PopupScreen "Comandos Perfiladores" 1280x714
   Button "Botón_6" at 630,585 size 88x33; TextOff 'Avance'
      on Press: SetTag("DB_OP.RC1", 52); SetBit("DB_OP.OP_SELMANU1")
      Visibility <- "MANU"
      Appearance <- "DB_OP.RC1"
   Button "Botón_7" at 630,630 size 88x33; TextOff 'Retroceso'
      on Press: SetTag("DB_OP.RC1", 53); SetBit("DB_OP.OP_SELMANU1")
      Visibility <- "MANU"
      Appearance <- "DB_OP.RC1"
   Button "Botón_8" at 731,585 size 88x33; TextOff 'Hacia Consigna'
      on Press: SetTag("DB_OP.RC1", 51); SetBit("DB_OP.OP_SELMANU1")
      Visibility <- "MANU"
      Appearance <- "DB_OP.RC1"
   Button "Botón_11" at 731,630 size 88x33; TextOff 'Freno'
      on Press: SetTag("DB_OP.RC1", 54); SetBit("DB_OP.OP_SELMANU1")
      Visibility <- "MANU"
      Appearance <- "DB_OP.RC1"
   Button "Botón_1" at 889,270 size 88x33; TextOff 'Avance'
      on Press: SetTag("DB_OP.RC1", 55); SetBit("DB_OP.OP_SELMANU1")
      Visibility <- "MANU"
      Appearance <- "DB_OP.RC1"
   Button "Botón_2" at 889,307 size 88x33; TextOff 'Retroceso'
      on Press: SetTag("DB_OP.RC1", 56); SetBit("DB_OP.OP_SELMANU1")
      Visibility <- "MANU"
      Appearance <- "DB_OP.RC1"
   IOField "Champ E/S_1" at 943,573 size 77x29; FormatPattern 9999999
      ProcessValue <- "DB_OP.COD1_VAL"
   IOField "Champ E/S" at 947,636 size 70x29; FormatPattern 9.9999
      ProcessValue <- "DB_OP.COD1_COEF"
   IOField "Champ E/S_0" at 943,601 size 77x29; FormatPattern 9999999
      ProcessValue <- "DB_OP.COD1_CONS"
   IOField "Champ E/S_2" at 1114,575 size 69x29; FormatPattern 9999999
      ProcessValue <- "DB_OP.COD1_INIT"
   TextField "Champ de texte_2" at 861,578 size 82x18; Text 'Posición / Position Réelle'
   TextField "Champ de texte" at 844,607 size 99x18; Text 'Consigna / Position Consigne'
   TextField "Champ de texte_0" at 851,641 size 92x18; Text 'Coef corrección / Coeff correction'
   IOField "Champ E/S_4" at 1114,640 size 69x29; FormatPattern 9999999
      ProcessValue <- "DB_OP.COD1_TARGET"
   TextField "Champ de texte_5" at 1044,612 size 62x18; Text 'Cota Paro / Côte Arrêt'
   TextField "Champ de texte_6" at 1052,645 size 50x18; Text 'Ventana / Fenetre'
   IOField "Champ E/S_5" at 1114,607 size 69x29; FormatPattern 9999999
      ProcessValue <- "DB_OP.COD1_ARRET"
   Button "Button" at 1045,578 size 60x23; TextOff 'OFFSET'; Authorization "Nivel 1"
      on Press: SetBit("DB_OP.COD1_CMD")
      Appearance <- "DB_OP.COD2_CMD"
   GraphicIOField "Campo ES gráfico_4" at 236,203 size 456x232; PictureList "Grupo 2 - Perfilador"
      ProcessValue <- "Alarma_Perfiladores"
   Polygon "Polígono_3" at 265,240 size 389x46
      Visibility <- "Perfiladores\Perfilador.PresenciaPieza"
   Rectangle "Rectángulo_2" at 874,227 size 118x128
      Visibility <- "MANU"
   Rectangle "Rectángulo_3" at 874,227 size 118x29
      Visibility <- "MANU"
   TextField "Campo de texto_1" at 900,231 size 66x18; Text 'Perfiladores'
      Visibility <- "MANU"
   Circle "Cercle_11" at 450,253 size 12x12
      Appearance <- "27S4"
   Circle "Cercle_12" at 413,405 size 12x12
      Appearance <- "29S7"
   Circle "Cercle_13" at 411,387 size 12x12
      Appearance <- "29S7"
   Circle "Cercle_14" at 515,384 size 12x12
      Appearance <- "23S4"
   Polygon "Polígono_1" at 248,269 size 17x19
      Appearance <- "36S70"
   TextField "Campo de texto_3" at 246,143 size 112x18; Text 'Sensores de Atasco'
   TextField "Campo de texto_4" at 613,454 size 141x18; Text '23S4 - Presión de Frenos'
   TextField "Campo de texto_5" at 414,107 size 101x18; Text 'Motor Perfilador 4'
   TextField "Campo de texto_6" at 684,429 size 101x18; Text 'Motor Perfilador 3'
   TextField "Campo de texto_7" at 159,441 size 101x18; Text 'Motor Perfilador 1'
   TextField "Campo de texto_8" at 147,165 size 101x18; Text 'Motor Perfilador 2'
   TextField "Campo de texto_9" at 140,188 size 64x46; Text '36S70 Barrera de Atascos'
   TextField "Campo de texto_10" at 557,500 size 197x18; Text 'M07 - Motor Ajuste de Profundidad'
   TextField "Campo de texto_11" at 202,476 size 119x18; Text '29S7 - Fin de Carrera'
   TextField "Campo de texto_13" at 320,502 size 53x18; Text 'Encóder'
   TextField "Campo de texto_14" at 118,363 size 81x46; Text '27S3 - Chapa en Entrada Perfilador'
   Circle "Cercle_2" at 236,274 size 12x12
      Appearance <- "27S3"
   Polyline "Línea poligonal_11" at 263,255 size 397x22
      Appearance <- "36S70"
   Polygon "Polígono_2" at 655,246 size 17x19
      Appearance <- "36S70"
   Rectangle "Rectángulo_6" at 613,555 size 222x128
      Visibility <- "MANU"
   Rectangle "Rectángulo_7" at 834,539 size 374x144
      Visibility <- "MANU"
   Rectangle "Rectángulo_8" at 613,539 size 595x29
      Visibility <- "MANU"
   TextField "Campo de texto_12" at 674,543 size 108x18; Text 'Ajuste Profundidad'
      Visibility <- "MANU"

PopupScreen "Comandos Cinta" 1280x714
   Button "Botón_6" at 630,585 size 88x33; TextOff 'Avance'
      on Press: SetTag("DB_OP.RC1", 52); SetBit("DB_OP.OP_SELMANU1")
      Visibility <- "MANU"
      Appearance <- "DB_OP.RC1"
   Button "Botón_7" at 630,630 size 88x33; TextOff 'Retroceso'
      on Press: SetTag("DB_OP.RC1", 53); SetBit("DB_OP.OP_SELMANU1")
      Visibility <- "MANU"
      Appearance <- "DB_OP.RC1"
   Button "Botón_8" at 731,585 size 88x33; TextOff 'Hacia Consigna'
      on Press: SetTag("DB_OP.RC1", 51); SetBit("DB_OP.OP_SELMANU1")
      Visibility <- "MANU"
      Appearance <- "DB_OP.RC1"
   Button "Botón_11" at 731,630 size 88x33; TextOff 'Freno'
      on Press: SetTag("DB_OP.RC1", 54); SetBit("DB_OP.OP_SELMANU1")
      Visibility <- "MANU"
      Appearance <- "DB_OP.RC1"
   Button "Botón_4" at 462,582 size 88x33; TextOff 'Avance'
      on Press: SetTag("DB_OP.RC2", 91); SetBit("DB_OP.OP_SELMANU2")
      Visibility <- "MANU"
      Appearance <- "DB_OP.RC2"
   Button "Botón_5" at 462,619 size 88x33; TextOff 'Retroceso'
      on Press: SetTag("DB_OP.RC2", 92); SetBit("DB_OP.OP_SELMANU2")
      Visibility <- "MANU"
      Appearance <- "DB_OP.RC2"
   IOField "Champ E/S_1" at 943,573 size 77x29; FormatPattern 9999999
      ProcessValue <- "DB_OP.COD2_VAL"
   IOField "Champ E/S" at 947,636 size 70x29; FormatPattern 9.9999
      ProcessValue <- "DB_OP.COD2_COEF"
   IOField "Champ E/S_0" at 943,601 size 77x29; FormatPattern 9999999
      ProcessValue <- "DB_OP.COD2_CONS"
   IOField "Champ E/S_2" at 1114,575 size 69x29; FormatPattern 9999999
      ProcessValue <- "DB_OP.COD2_INIT"
   TextField "Champ de texte_2" at 861,578 size 82x18; Text 'Posición / Position Réelle'
   TextField "Champ de texte" at 844,607 size 99x18; Text 'Consigna / Position Consigne'
   TextField "Champ de texte_0" at 851,641 size 92x18; Text 'Coef corrección / Coeff correction'
   IOField "Champ E/S_4" at 1114,640 size 69x29; FormatPattern 9999999
      ProcessValue <- "DB_OP.COD2_TARGET"
   TextField "Champ de texte_5" at 1044,612 size 62x18; Text 'Cota Paro / Côte Arrêt'
   TextField "Champ de texte_6" at 1052,645 size 50x18; Text 'Ventana / Fenetre'
   IOField "Champ E/S_5" at 1114,607 size 69x29; FormatPattern 9999999
      ProcessValue <- "DB_OP.COD2_ARRET"
   Button "Button" at 1045,578 size 60x23; TextOff 'OFFSET'; Authorization "Nivel 1"
      on Press: SetBit("DB_OP.COD2_CMD")
      Appearance <- "DB_OP.COD2_CMD"
   GraphicIOField "Campo ES gráfico_1" at 290,222 size 647x180; PictureList "Grupo 2 - Cinta"
      ProcessValue <- "Alarma_Cinta"
   Rectangle "Rectángulo_1" at 613,555 size 222x128
      Visibility <- "MANU"
   Rectangle "Rectángulo_2" at 448,539 size 118x128
      Visibility <- "MANU"
   Rectangle "Rectángulo_3" at 448,539 size 118x29
      Visibility <- "MANU"
   TextField "Campo de texto_1" at 474,543 size 31x18; Text 'Cinta'
      Visibility <- "MANU"
   Rectangle "Rectángulo_6" at 834,539 size 374x144
      Visibility <- "MANU"
   Rectangle "Rectángulo_7" at 613,539 size 595x29
      Visibility <- "MANU"
   TextField "Campo de texto_12" at 642,543 size 108x18; Text 'Ajuste Profundidad'
      Visibility <- "MANU"
   Circle "Cercle_1" at 325,248 size 12x12
      Appearance <- "27S4"
   Circle "Cercle_14" at 909,220 size 12x12
      Appearance <- "29S1"
   Circle "Cercle_15" at 909,234 size 12x12
      Appearance <- "29S2"
   Circle "Cercle_11" at 826,289 size 12x12
      Appearance <- "25S2"
   Circle "Cercle" at 911,284 size 12x12
      Appearance <- "29S3"
   TextField "Campo de texto_22" at 109,219 size 183x18; Text '27S4 - Chapa en Salida Perfilador'
   TextField "Campo de texto_23" at 624,433 size 179x18; Text 'M07 - Motor Ajuste Profundidad'
   TextField "Campo de texto_24" at 987,328 size 126x18; Text '25S2 - Bajar Velocidad'
   TextField "Campo de texto_25" at 512,385 size 223x18; Text '29S3 - Presencia de Chapa en Formador'
   TextField "Campo de texto_31" at 616,197 size 166x18; Text 'M08 - Motor Transporte Cinta'
   TextField "Campo de texto_32" at 667,130 size 145x18; Text '29S1 - Avance Bloqueado'
   TextField "Campo de texto_33" at 647,164 size 165x18; Text '29S2 - Avance Desbloqueado'
   Polygon "Polígono_4" at 351,252 size 385x62
      Visibility <- "Cinta\Cinta.PresenciaPieza"

PopupScreen "Comandos Descargador" 1280x714
   GraphicView "Visor de gráficos_1" at 134,166 size 538x272; Picture "Rolos 3"
   Rectangle "Rectángulo_9" at 811,197 size 118x128
      Visibility <- "MANU"
   Rectangle "Rectángulo_8" at 811,197 size 118x29
      Visibility <- "MANU"
   TextField "Campo de texto_3" at 854,201 size 32x18; Text 'Rolos'
      Visibility <- "MANU"
   Button "Botón_29" at 826,241 size 88x33; TextOff 'Avance'
      on Press: SetTag("DB_OP.RC1", 41); SetBit("DB_OP.OP_SELMANU1")
      Visibility <- "MANU"
      Appearance <- "DB_OP.RC1"
   Button "Botón_30" at 826,279 size 88x33; TextOff 'Retroceso'
      on Press: SetTag("DB_OP.RC1", 42); SetBit("DB_OP.OP_SELMANU1")
      Visibility <- "MANU"
      Appearance <- "DB_OP.RC1"
   TextField "Campo de texto_7" at 303,476 size 104x32; Text '27S3 - Chapa en Entrada Perfilador'
   Circle "Cercle_10" at 201,328 size 12x12
      Appearance <- "27S3"
   Circle "Cercle_13" at 349,283 size 12x12
      Appearance <- "26S8"
   TextField "Campo de texto_11" at 455,437 size 114x32; Text '26S8 - Chapa en Transporte de Rolos'

screen "eProC - 01 Araña" 1280x768, template "Template"
   Polygon "Polígono_3" at 343,318 size 325x50
      Visibility <- "Araña\Araña.PresenciaPieza"
   Rectangle "Rectángulo_7" at 989,250 size 248x208
      Visibility <- "MANU"
   Rectangle "Rectángulo_12" at 989,246 size 248x29
      Visibility <- "MANU"
   Rectangle "Rectángulo_9" at 843,563 size 118x128
      Visibility <- "MANU"
   Rectangle "Rectángulo_8" at 843,563 size 118x29
      Visibility <- "MANU"
   TextField "Campo de texto_3" at 870,567 size 64x18; Text 'Transporte'
      Visibility <- "MANU"
   TextField "Campo de texto_11" at 1010,252 size 66x18; Text 'Aire Tulipas'
      Visibility <- "MANU"
   Button "Botón_4" at 859,607 size 88x33; TextOff 'Avance'
      on Press: SetTag("DB_OP.RC1", 11); SetBit("DB_OP.OP_SELMANU1")
      Visibility <- "MANU"
      Appearance <- "DB_OP.RC1"
   Button "Botón_5" at 859,645 size 88x33; TextOff 'Retroceso'
      on Press: SetTag("DB_OP.RC1", 12); SetBit("DB_OP.OP_SELMANU1")
      Visibility <- "MANU"
      Appearance <- "DB_OP.RC1"
   Button "Botón_10" at 1065,290 size 72x33; TextOff 'Activar'
      on Press: SetTag("DB_OP.RC1", 20); SetBit("DB_OP.OP_SELMANU1")
      Visibility <- "MANU"
      Appearance <- "DB_OP.RC1"
   Button "Botón_17" at 1145,290 size 72x33; TextOff 'Desactivar'
      on Press: SetTag("DB_OP.RC1", 21); SetBit("DB_OP.OP_SELMANU1")
      Visibility <- "MANU"
      Appearance <- "DB_OP.RC1"
   TextField "Campo de texto_12" at 1010,296 size 37x18; Text 'Todas'
      Visibility <- "MANU"
   Button "Botón_1" at 1065,336 size 72x33; TextOff 'Activar'
      on Press: SetTag("DB_OP.RC1", 32); SetBit("DB_OP.OP_SELMANU1")
      Visibility <- "MANU"
      Appearance <- "DB_OP.RC1"
   Button "Botón_23" at 1065,373 size 72x33; TextOff 'Activar'
      on Press: SetTag("DB_OP.RC1", 34); SetBit("DB_OP.OP_SELMANU1")
      Visibility <- "MANU"
      Appearance <- "DB_OP.RC1"
   Button "Botón_24" at 1065,411 size 72x33; TextOff 'Activar'
      on Press: SetTag("DB_OP.RC1", 36); SetBit("DB_OP.OP_SELMANU1")
      Visibility <- "MANU"
      Appearance <- "DB_OP.RC1"
   Button "Botón_26" at 1145,336 size 72x33; TextOff 'Desactivar'
      on Press: SetTag("DB_OP.RC1", 33); SetBit("DB_OP.OP_SELMANU1")
      Visibility <- "MANU"
      Appearance <- "DB_OP.RC1"
   Button "Botón_27" at 1145,373 size 72x33; TextOff 'Desactivar'
      on Press: SetTag("DB_OP.RC1", 35); SetBit("DB_OP.OP_SELMANU1")
      Visibility <- "MANU"
      Appearance <- "DB_OP.RC1"
   Button "Botón_28" at 1145,411 size 72x33; TextOff 'Desactivar'
      on Press: SetTag("DB_OP.RC1", 37); SetBit("DB_OP.OP_SELMANU1")
      Visibility <- "MANU"
      Appearance <- "DB_OP.RC1"
   TextField "Campo de texto_2" at 1008,343 size 48x18; Text 'Grupo 1'
      Visibility <- "MANU"
   TextField "Campo de texto_1" at 1008,381 size 48x18; Text 'Grupo 2'
      Visibility <- "MANU"
   TextField "Campo de texto_5" at 1008,419 size 48x18; Text 'Grupo 3'
      Visibility <- "MANU"
   Rectangle "Rectángulo_1" at 989,483 size 248x208
      Visibility <- "MANU"
   Rectangle "Rectángulo_2" at 989,479 size 248x29
      Visibility <- "MANU"
   TextField "Campo de texto_13" at 1010,485 size 74x18; Text 'Vacío Tulipas'
      Visibility <- "MANU"
   TextField "Campo de texto_14" at 1010,529 size 37x18; Text 'Todas'
      Visibility <- "MANU"
   TextField "Campo de texto_15" at 1008,576 size 48x18; Text 'Grupo 1'
      Visibility <- "MANU"
   TextField "Campo de texto_16" at 1008,614 size 48x18; Text 'Grupo 2'
      Visibility <- "MANU"
   TextField "Campo de texto_17" at 1008,652 size 48x18; Text 'Grupo 3'
      Visibility <- "MANU"
   Button "Botón_21" at 1065,523 size 72x33; TextOff 'Activar'
      on Press: SetTag("DB_OP.RC1", 30); SetBit("DB_OP.OP_SELMANU1")
      Visibility <- "MANU"
      Appearance <- "DB_OP.RC1"
   Button "Botón_25" at 1145,523 size 72x33; TextOff 'Desactivar'
      on Press: SetTag("DB_OP.RC1", 31); SetBit("DB_OP.OP_SELMANU1")
      Visibility <- "MANU"
      Appearance <- "DB_OP.RC1"
   Button "Botón_14" at 1065,569 size 72x33; TextOff 'Activar'
      on Press: SetTag("DB_OP.RC1", 22); SetBit("DB_OP.OP_SELMANU1")
      Visibility <- "MANU"
      Appearance <- "DB_OP.RC1"
   Button "Botón_15" at 1065,606 size 72x33; TextOff 'Activar'
      on Press: SetTag("DB_OP.RC1", 24); SetBit("DB_OP.OP_SELMANU1")
      Visibility <- "MANU"
      Appearance <- "DB_OP.RC1"
   Button "Botón_16" at 1065,644 size 72x33; TextOff 'Activar'
      on Press: SetTag("DB_OP.RC1", 26); SetBit("DB_OP.OP_SELMANU1")
      Visibility <- "MANU"
      Appearance <- "DB_OP.RC1"
   Button "Botón_18" at 1145,569 size 72x33; TextOff 'Desactivar'
      on Press: SetTag("DB_OP.RC1", 23); SetBit("DB_OP.OP_SELMANU1")
      Visibility <- "MANU"
      Appearance <- "DB_OP.RC1"
   Button "Botón_19" at 1145,606 size 72x33; TextOff 'Desactivar'
      on Press: SetTag("DB_OP.RC1", 25); SetBit("DB_OP.OP_SELMANU1")
      Visibility <- "MANU"
      Appearance <- "DB_OP.RC1"
   Button "Botón_20" at 1145,644 size 72x33; TextOff 'Desactivar'
      on Press: SetTag("DB_OP.RC1", 27); SetBit("DB_OP.OP_SELMANU1")
      Visibility <- "MANU"
      Appearance <- "DB_OP.RC1"
   Rectangle "Rectángulo_10" at 988,26 size 248x201
      Visibility <- "MANU"
   Button "Botón_6" at 1012,65 size 202x33; TextOff 'Subir (Pistón Superior)'
      on Press: SetTag("DB_OP.RC1", 16); SetBit("DB_OP.OP_SELMANU1")
      Visibility <- "MANU"
      Appearance <- "DB_OP.RC1"
   Button "Botón_7" at 1012,103 size 202x33; TextOff 'Bajar (Pistón Superior)'
      on Press: SetTag("DB_OP.RC1", 15); SetBit("DB_OP.OP_SELMANU1")
      Visibility <- "MANU"
      Appearance <- "DB_OP.RC1"
   Button "Botón_8" at 1012,179 size 202x33; TextOff 'Bajar (Pistón Inferior)'
      on Press: SetTag("DB_OP.RC1", 13); SetBit("DB_OP.OP_SELMANU1")
      Visibility <- "MANU"
      Appearance <- "DB_OP.RC1"
   Button "Botón_9" at 1012,141 size 202x33; TextOff 'Subir (Pistón Inferior)'
      on Press: SetTag("DB_OP.RC1", 14); SetBit("DB_OP.OP_SELMANU1")
      Visibility <- "MANU"
      Appearance <- "DB_OP.RC1"
   Rectangle "Rectángulo_11" at 988,26 size 248x29
      Visibility <- "MANU"
   TextField "Campo de texto_7" at 1056,30 size 110x18; Text 'Movimiento Vertical'
      Visibility <- "MANU"
   GraphicIOField "Campo ES gráfico_1" at 295,98 size 460x334; PictureList "Araña"
      ProcessValue <- "Alarma_Araña"
   Button "Botón_2" at 453,467 size 144x49; TextOff 'Inicializar'
      on Press: SetBit("Comando_Inicializar_Araña")
      Visibility <- "MANU"
   Group "Group" at 428,460 size 189x68
   TextField "Campo de texto_8" at 61,77 size 35x18; Text 'Araña'
   TextField "Campo de texto_18" at 61,98 size 12x18; Text 'A'
   IOField "Champ E/S_8" at 98,95 size 54x25; FormatPattern 9999999
      Appearance <- "Araña\Araña.PresenciaPieza"
      ProcessValue <- "Araña\Araña.A"
   IOField "Champ E/S_9" at 98,115 size 54x25; FormatPattern 9999999
      Appearance <- "Araña\Araña.PresenciaPieza"
      ProcessValue <- "Araña\Araña.B"
   IOField "Champ E/S_10" at 98,136 size 54x24; FormatPattern 9999999
      Appearance <- "Araña\Araña.PresenciaPieza"
      ProcessValue <- "Araña\Araña.C"
   IOField "Champ E/S_11" at 98,155 size 54x25; FormatPattern 9999999
      Appearance <- "Araña\Araña.PresenciaPieza"
      ProcessValue <- "Araña\Araña.D"
   TextField "Campo de texto_29" at 62,116 size 11x18; Text 'B'
   TextField "Campo de texto_30" at 62,136 size 11x18; Text 'C'
   TextField "Campo de texto_31" at 62,156 size 12x18; Text 'D'
   Button "Botón_3" at 45,40 size 128x33; TextOff 'Borrar Pieza'
      on Click: ResetBit("Araña\Araña.PresenciaPieza")
      Visibility <- "Araña\Araña.PresenciaPieza"
   Button "Botón_12" at 45,340 size 128x33; TextOff 'Transferir Datos'
      on Click: SetBit("Forz_Transf1")
      Visibility <- "Perfiladores\Perfilador.PresenciaPieza"
   Button "Template_Plantilla_Botón_3" at 1,688 size 130x29; TextOff 'ARAÑA'
   Button "Plantilla_Botón_1" at 1,715 size 130x53; TextOff 'PRINCIPAL'
      on Click: ActivateScreen("eProC - Principal", 0)
   Button "Template_Plantilla_Bouton_2" at 1085,715 size 193x53; TextOff 'ALARMAS / DEFAUT'
      on Press: ActivateScreen("eProC - Alarmas", 0)
      Visibility <- "DB_OP.P_DEFAUT"
   Circle "Cercle_11" at 494,226 size 10x10
      Appearance <- "25S8"
   Circle "Cercle_12" at 495,183 size 10x10
      Appearance <- "25S7"
   Circle "Cercle_0" at 494,247 size 10x10
      Appearance <- "25S4"
   Circle "Cercle_1" at 534,134 size 10x10
      Appearance <- "25S3"
   Circle "Cercle_2" at 538,186 size 10x10
      Appearance <- "25S5"
   TextField "Campo de texto_6" at 645,56 size 186x22; Text '25S3 - Fin de Carrera Arriba'
   TextField "Campo de texto_9" at 620,126 size 186x22; Text '25S5 - Fin de Carrera Abajo'
   TextField "Campo de texto_19" at 218,103 size 174x22; Text '25S7 - Pistón 2 Expandido'
   TextField "Campo de texto_20" at 220,139 size 169x22; Text '25S8 - Pistón 2 Contraído'
   TextField "Campo de texto_21" at 220,198 size 169x22; Text '25S4 - Pistón 1 Contraído'
   TextField "Campo de texto_22" at 297,228 size 132x22; Text '25S6 - Araña Abajo'
   Circle "Cercle_5" at 457,251 size 10x10
      Appearance <- "25S6"
   Circle "Cercle" at 476,339 size 10x10
      Appearance <- "26S1"
   TextField "Campo de texto_23" at 183,430 size 248x22; Text '26S1 - Tulipas Apoyadas en la Chapa'
   TextField "Campo de texto_24" at 768,228 size 151x22; Text '26S5 - Bajar Velocidad'
   TextField "Campo de texto_25" at 763,204 size 210x22; Text '26S3 - En Posición de Descarga'
   TextField "Campo de texto_26" at 773,293 size 206x58; Text 'M03 - Motor Transporte Araña KM02.1 -> Hacia Rolos KM02.2 -> Hacia Almacenes'
   TextField "Campo de texto_27" at 785,393 size 151x22; Text '26S4 - Bajar Velocidad'
   TextField "Campo de texto_28" at 787,418 size 187x22; Text '26S2 - En Posición de Carga'
   Circle "Cercle_4" at 701,406 size 10x10
      Appearance <- "26S2"
   Circle "Cercle_6" at 696,382 size 10x10
      Appearance <- "26S4"
   Circle "Cercle_7" at 681,214 size 10x10
      Appearance <- "26S5"
   Circle "Cercle_8" at 676,191 size 10x10
      Appearance <- "26S3"
   Rectangle "Rectángulo_3" at 428,460 size 189x68
      Visibility <- "Araña_Inicializada"
   TextField "Campo de texto_4" at 442,481 size 159x22; Text 'Araña en Posición Inicial'
      Visibility <- "Araña_Inicializada"
   TextField "Campo de texto_142" at 62,178 size 17x18; Text 'F1'
   IOField "Champ E/S_134" at 102,175 size 51x25; FormatPattern s999999
      Appearance <- "Araña\Araña.PresenciaPieza"
      ProcessValue <- "Araña\Araña.F1"
   IOField "Champ E/S_135" at 102,195 size 51x25; FormatPattern s999999
      Appearance <- "Araña\Araña.PresenciaPieza"
      ProcessValue <- "Araña\Araña.F2"
   IOField "Champ E/S_136" at 102,216 size 51x24; FormatPattern s999999
      Appearance <- "Araña\Araña.PresenciaPieza"
      ProcessValue <- "Araña\Araña.F3"
   IOField "Champ E/S_137" at 102,235 size 51x25; FormatPattern s999999
      Appearance <- "Araña\Araña.PresenciaPieza"
      ProcessValue <- "Araña\Araña.F4"
   TextField "Campo de texto_143" at 62,197 size 17x18; Text 'F2'
   TextField "Campo de texto_144" at 62,217 size 17x18; Text 'F3'
   TextField "Campo de texto_145" at 62,237 size 17x18; Text 'F4'
   TextField "Campo de texto_146" at 62,258 size 35x18; Text 'PL1-1'
   IOField "Champ E/S_138" at 102,255 size 51x25; FormatPattern s999999
      Appearance <- "Araña\Araña.PresenciaPieza"
      ProcessValue <- "Araña\Araña.PL1_1"
   IOField "Champ E/S_139" at 102,275 size 51x25; FormatPattern s999999
      Appearance <- "Araña\Araña.PresenciaPieza"
      ProcessValue <- "Araña\Araña.PL1_2"
   IOField "Champ E/S_140" at 102,296 size 51x24; FormatPattern s999999
      Appearance <- "Araña\Araña.PresenciaPieza"
      ProcessValue <- "Araña\Araña.PL2_1"
   IOField "Champ E/S_141" at 102,315 size 51x25; FormatPattern s999999
      Appearance <- "Araña\Araña.PresenciaPieza"
      ProcessValue <- "Araña\Araña.PL2_2"
   TextField "Campo de texto_147" at 62,278 size 35x18; Text 'PL1-2'
   TextField "Campo de texto_148" at 62,299 size 35x18; Text 'PL2-1'
   TextField "Campo de texto_149" at 62,318 size 35x18; Text 'PL2-2'

screen "eProC - 02 Rolos" 1280x768, template "Template"
   GraphicIOField "Campo ES gráfico_4" at 286,166 size 538x272; PictureList "Rolos"
      ProcessValue <- "Alarma_Perfiladores"
   Polygon "Polígono_3" at 336,215 size 385x136
      Visibility <- "Rolos\Rolos.PresenciaPieza"
   Rectangle "Rectángulo_9" at 963,197 size 118x128
      Visibility <- "MANU"
   Rectangle "Rectángulo_8" at 963,197 size 118x29
      Visibility <- "MANU"
   TextField "Campo de texto_3" at 1006,201 size 32x18; Text 'Rolos'
      Visibility <- "MANU"
   Button "Botón_29" at 978,241 size 88x33; TextOff 'Avance'
      on Press: SetTag("DB_OP.RC1", 41); SetBit("DB_OP.OP_SELMANU1")
      Visibility <- "MANU"
      Appearance <- "DB_OP.RC1"
   Button "Botón_30" at 978,279 size 88x33; TextOff 'Retroceso'
      on Press: SetTag("DB_OP.RC1", 42); SetBit("DB_OP.OP_SELMANU1")
      Visibility <- "MANU"
      Appearance <- "DB_OP.RC1"
   TextField "Campo de texto_7" at 455,476 size 124x40; Text '27S3 - Chapa en Entrada Perfilador'
   Circle "Cercle_10" at 353,328 size 12x12
      Appearance <- "27S3"
   Circle "Cercle_13" at 613,248 size 12x12
      Appearance <- "26S8"
   TextField "Campo de texto_11" at 719,402 size 137x40; Text '26S8 - Chapa en Transporte de Rolos'
   TextField "Campo de texto_10" at 61,77 size 32x18; Text 'Rolos'
   TextField "Campo de texto_20" at 61,99 size 12x18; Text 'A'
   IOField "Champ E/S_12" at 96,95 size 54x25; FormatPattern 9999999
      Appearance <- "Rolos\Rolos.PresenciaPieza"
      ProcessValue <- "Rolos\Rolos.A"
   IOField "Champ E/S_13" at 96,115 size 54x25; FormatPattern 9999999
      Appearance <- "Rolos\Rolos.PresenciaPieza"
      ProcessValue <- "Rolos\Rolos.B"
   IOField "Champ E/S_14" at 96,136 size 54x24; FormatPattern 9999999
      Appearance <- "Rolos\Rolos.PresenciaPieza"
      ProcessValue <- "Rolos\Rolos.C"
   IOField "Champ E/S_15" at 96,155 size 54x25; FormatPattern 9999999
      Appearance <- "Rolos\Rolos.PresenciaPieza"
      ProcessValue <- "Rolos\Rolos.D"
   TextField "Campo de texto_21" at 61,117 size 11x18; Text 'B'
   TextField "Campo de texto_22" at 61,137 size 11x18; Text 'C'
   TextField "Campo de texto_23" at 61,157 size 12x18; Text 'D'
   Button "Botón_9" at 45,40 size 126x33; TextOff 'Borrar Pieza'
      on Click: ResetBit("Rolos\Rolos.PresenciaPieza")
      Visibility <- "Rolos\Rolos.PresenciaPieza"
   Button "Botón_4" at 45,340 size 128x33; TextOff 'Transferir Datos'
      on Click: SetBit("Forz_Transf2")
      Visibility <- "Perfiladores\Perfilador.PresenciaPieza"
   Button "Template_Plantilla_Botón_3" at 1,688 size 130x29; TextOff 'ROLOS'
   Button "Plantilla_Botón_1" at 1,715 size 130x53; TextOff 'PRINCIPAL'
      on Click: ActivateScreen("eProC - Principal", 0)
   Button "Template_Plantilla_Bouton_2" at 1085,715 size 193x53; TextOff 'ALARMAS / DEFAUT'
      on Press: ActivateScreen("eProC - Alarmas", 0)
      Visibility <- "DB_OP.P_DEFAUT"
   TextField "Campo de texto_134" at 62,178 size 17x18; Text 'F1'
   IOField "Champ E/S_126" at 102,175 size 51x25; FormatPattern s999999
      Appearance <- "Rolos\Rolos.PresenciaPieza"
      ProcessValue <- "Rolos\Rolos.F1"
   IOField "Champ E/S_127" at 102,195 size 51x25; FormatPattern s999999
      Appearance <- "Rolos\Rolos.PresenciaPieza"
      ProcessValue <- "Rolos\Rolos.F2"
   IOField "Champ E/S_128" at 102,216 size 51x24; FormatPattern s999999
      Appearance <- "Rolos\Rolos.PresenciaPieza"
      ProcessValue <- "Rolos\Rolos.F3"
   IOField "Champ E/S_129" at 102,235 size 51x25; FormatPattern s999999
      Appearance <- "Rolos\Rolos.PresenciaPieza"
      ProcessValue <- "Rolos\Rolos.F4"
   TextField "Campo de texto_135" at 62,197 size 17x18; Text 'F2'
   TextField "Campo de texto_136" at 62,217 size 17x18; Text 'F3'
   TextField "Campo de texto_137" at 62,237 size 17x18; Text 'F4'
   TextField "Campo de texto_138" at 62,258 size 35x18; Text 'PL1-1'
   IOField "Champ E/S_130" at 102,255 size 51x25; FormatPattern s999999
      Appearance <- "Rolos\Rolos.PresenciaPieza"
      ProcessValue <- "Rolos\Rolos.PL1_1"
   IOField "Champ E/S_131" at 102,275 size 51x25; FormatPattern s999999
      Appearance <- "Rolos\Rolos.PresenciaPieza"
      ProcessValue <- "Rolos\Rolos.PL1_2"
   IOField "Champ E/S_132" at 102,296 size 51x24; FormatPattern s999999
      Appearance <- "Rolos\Rolos.PresenciaPieza"
      ProcessValue <- "Rolos\Rolos.PL2_1"
   IOField "Champ E/S_133" at 102,315 size 51x25; FormatPattern s999999
      Appearance <- "Rolos\Rolos.PresenciaPieza"
      ProcessValue <- "Rolos\Rolos.PL2_2"
   TextField "Campo de texto_139" at 62,278 size 35x18; Text 'PL1-2'
   TextField "Campo de texto_140" at 62,299 size 35x18; Text 'PL2-1'
   TextField "Campo de texto_141" at 62,318 size 35x18; Text 'PL2-2'

screen "eProC - 00 Almacenes" 1280x768, template "Template"
   Rectangle "Rectángulo_9" at 1020,194 size 118x128
      Visibility <- "MANU"
   Rectangle "Rectángulo_8" at 1020,194 size 118x29
      Visibility <- "MANU"
   TextField "Campo de texto_3" at 1036,198 size 86x18; Text 'Intercambiador'
      Visibility <- "MANU"
   Button "Botón_1" at 1035,238 size 88x33; TextOff 'Avance'
      on Press: SetTag("DB_OP.RC1", 1); SetBit("DB_OP.OP_SELMANU1")
      Visibility <- "MANU"
      Appearance <- "DB_OP.RC1"
   Button "Botón_2" at 1035,276 size 88x33; TextOff 'Retroceso'
      on Press: SetTag("DB_OP.RC1", 2); SetBit("DB_OP.OP_SELMANU1")
      Visibility <- "MANU"
      Appearance <- "DB_OP.RC1"
   TextField "Campo de texto_2" at 95,341 size 267x22; Text '26S7 - Almacén 2 en puesto de Trabajo'
   TextField "Campo de texto_4" at 175,412 size 260x22; Text '26S6 - Almacén 2 en puesto de Espera'
   GraphicIOField "Campo ES gráfico_2" at 480,113 size 396x294; PictureList "Grupo 1 - Almacén A"
      ProcessValue <- "26S7"
   GraphicIOField "Campo ES gráfico_1" at 480,113 size 396x294; PictureList "Grupo 1 - Almacén B"
      ProcessValue <- "26S7"
      Visibility <- "Alarma_Almacenes"
   Circle "Cercle_2" at 486,298 size 14x14
      Appearance <- "26S7"
   TextField "Campo de texto_6" at 132,470 size 286x22; Text 'M01 - Motor Intercambiador de Almacenes'
   Circle "Cercle_1" at 565,354 size 14x14
      Appearance <- "26S6"
   Polyline "Línea poligonal_11" at 542,162 size 264x133
      Appearance <- "36S10"
   TextField "Campo de texto_1" at 114,231 size 251x22; Text '36S10 - Barrera Seguridad Almacenes'
   Button "Botón_4" at 806,409 size 144x49; TextOff 'Habilitar'
      on Press: SetBit("Hab_Almacenes")
   Rectangle "Rectángulo_3" at 781,402 size 189x68
      Visibility <- "Enclavamiento"
   TextField "Campo de texto_5" at 800,423 size 148x22; Text 'Almacenes Habilitados'
      Visibility <- "Enclavamiento"
   Polygon "Polígono_2" at 800,152 size 20x12
      Appearance <- "36S10"
   Polygon "Polígono_1" at 528,288 size 20x12
      Appearance <- "36S10"
   Button "Template_Plantilla_Botón_3" at 1,688 size 130x29; TextOff 'ALMACENES'
   Button "Plantilla_Botón_1" at 1,715 size 130x53; TextOff 'PRINCIPAL'
      on Click: ActivateScreen("eProC - Principal", 0)
   Button "Template_Plantilla_Bouton_2" at 1085,715 size 193x53; TextOff 'ALARMAS / DEFAUT'
      on Press: ActivateScreen("eProC - Alarmas", 0)
      Visibility <- "DB_OP.P_DEFAUT"

screen "eProC - 03 Perfilador" 1280x768, template "Template"
   GraphicIOField "Campo ES gráfico_4" at 412,155 size 456x232; PictureList "Grupo 2 - Perfilador"
      ProcessValue <- "Alarma_Perfiladores"
   Polygon "Polígono_3" at 441,192 size 389x46
      Visibility <- "Perfiladores\Perfilador.PresenciaPieza"
   Rectangle "Rectángulo_2" at 987,531 size 118x144
      Visibility <- "MANU"
   Rectangle "Rectángulo_3" at 987,531 size 118x29
      Visibility <- "MANU"
   TextField "Campo de texto_1" at 1013,535 size 66x18; Text 'Perfiladores'
      Visibility <- "MANU"
   Circle "Cercle_11" at 458,214 size 12x12
      Appearance <- "Sensor 1"
   Circle "Cercle_13" at 587,339 size 12x12
      Appearance <- "29S6"
   Circle "Cercle_14" at 635,352 size 12x12
      Appearance <- "23S4"
   Polygon "Polígono_1" at 424,221 size 17x19
      Appearance <- "36S70"
   TextField "Campo de texto_3" at 406,92 size 134x22; Text 'Sensores de Atasco'
   TextField "Campo de texto_4" at 691,478 size 168x22; Text '23S4 - Presión de Frenos'
   TextField "Campo de texto_5" at 574,57 size 120x22; Text 'Motor Perfilador 4'
   TextField "Campo de texto_6" at 860,381 size 120x22; Text 'Motor Perfilador 3'
   TextField "Campo de texto_7" at 313,391 size 120x22; Text 'Motor Perfilador 1'
   TextField "Campo de texto_8" at 303,116 size 120x22; Text 'Motor Perfilador 2'
   TextField "Campo de texto_9" at 331,141 size 79x58; Text '36S70 Barrera de Atascos'
   TextField "Campo de texto_10" at 733,452 size 234x22; Text 'M07 - Motor Ajuste de Profundidad'
   TextField "Campo de texto_11" at 252,426 size 245x22; Text '29S6 - Fin de Carrera Hacia Adelante'
   TextField "Campo de texto_13" at 496,454 size 62x22; Text 'Encóder'
   TextField "Campo de texto_14" at 278,312 size 98x58; Text '27S3 - Chapa en Entrada Perfilador'
   Circle "Cercle_2" at 412,226 size 12x12
      Appearance <- "27S3"
   Polyline "Línea poligonal_11" at 439,207 size 397x22
      Appearance <- "36S70"
   Polygon "Polígono_2" at 831,198 size 17x19
      Appearance <- "36S70"
   Rectangle "Rectángulo_6" at 357,547 size 222x128
      Visibility <- "MANU"
   Rectangle "Rectángulo_8" at 357,531 size 222x29
      Visibility <- "MANU"
   TextField "Campo de texto_12" at 418,535 size 108x18; Text 'Ajuste Profundidad'
      Visibility <- "MANU"
   TextField "Campo de texto_2" at 61,77 size 54x18; Text 'Perfilador'
   TextField "Campo de texto_24" at 61,99 size 12x18; Text 'A'
   IOField "Champ E/S_16" at 100,95 size 53x25; FormatPattern 9999999
      Appearance <- "Perfiladores\Perfilador.PresenciaPieza"
      ProcessValue <- "Perfiladores\Perfilador.A"
   IOField "Champ E/S_17" at 100,115 size 53x25; FormatPattern 9999999
      Appearance <- "Perfiladores\Perfilador.PresenciaPieza"
      ProcessValue <- "Perfiladores\Perfilador.B"
   IOField "Champ E/S_18" at 100,136 size 53x24; FormatPattern 9999999
      Appearance <- "Perfiladores\Perfilador.PresenciaPieza"
      ProcessValue <- "Perfiladores\Perfilador.C"
   IOField "Champ E/S_19" at 100,155 size 53x25; FormatPattern 9999999
      Appearance <- "Perfiladores\Perfilador.PresenciaPieza"
      ProcessValue <- "Perfiladores\Perfilador.D"
   TextField "Campo de texto_25" at 63,117 size 11x18; Text 'B'
   TextField "Campo de texto_26" at 63,137 size 11x18; Text 'C'
   TextField "Campo de texto_27" at 63,157 size 12x18; Text 'D'
   Button "Botón_3" at 45,40 size 128x33; TextOff 'Borrar Pieza'
      on Click: ResetBit("Perfiladores\Perfilador.PresenciaPieza")
      Visibility <- "Perfiladores\Perfilador.PresenciaPieza"
   TextField "Campo de texto_16" at 754,420 size 232x22; Text '29S7 - Fin de Carrera Hacia Afuera'
   Circle "Cercle_3" at 696,349 size 12x12
      Appearance <- "29S7"
   Button "Botón_4" at 45,340 size 128x33; TextOff 'Transferir Datos'
      on Click: SetBit("Forz_Transf-3")
      Visibility <- "Perfiladores\Perfilador.PresenciaPieza"
   Circle "Cercle_4" at 474,213 size 12x12
      Appearance <- "Sensor 2"
   Circle "Cercle_5" at 490,211 size 12x12
      Appearance <- "Sensor 3"
   Circle "Cercle_6" at 506,210 size 12x12
      Appearance <- "Sensor 4"
   Circle "Cercle_7" at 522,209 size 12x12
      Appearance <- "Sensor 5"
   Circle "Cercle_8" at 538,208 size 12x12
      Appearance <- "Sensor 6"
   Circle "Cercle_9" at 554,207 size 12x12
      Appearance <- "Sensor 7"
   Circle "Cercle_10" at 570,206 size 12x12
      Appearance <- "Sensor 8"
   Circle "Cercle_12" at 586,205 size 12x12
      Appearance <- "Sensor 9"
   Circle "Cercle_15" at 602,203 size 12x12
      Appearance <- "Sensor 10"
   Circle "Cercle_16" at 618,202 size 12x12
      Appearance <- "Sensor 11"
   Circle "Cercle_17" at 634,201 size 12x12
      Appearance <- "Sensor 12"
   Circle "Cercle_18" at 650,200 size 12x12
      Appearance <- "Sensor 13"
   Circle "Cercle_19" at 666,199 size 12x12
      Appearance <- "Sensor 14"
   Circle "Cercle_20" at 682,198 size 12x12
      Appearance <- "Sensor 15"
   Circle "Cercle_21" at 698,197 size 12x12
      Appearance <- "Sensor 16"
   Circle "Cercle_22" at 714,196 size 12x12
      Appearance <- "Sensor 17"
   Circle "Cercle_23" at 730,195 size 12x12
      Appearance <- "Sensor 18"
   Circle "Cercle_24" at 746,194 size 12x12
      Appearance <- "Sensor 19"
   Circle "Cercle_25" at 762,193 size 12x12
      Appearance <- "Sensor 21"
   Circle "Cercle_26" at 778,192 size 12x12
      Appearance <- "Sensor 22"
   Circle "Cercle_27" at 794,191 size 12x12
      Appearance <- "Sensor 23"
   Circle "Cercle_28" at 810,190 size 12x12
      Appearance <- "Sensor 24"
   Button "Template_Plantilla_Botón_3" at 1,688 size 130x29; TextOff 'PERFILADOR'
   Button "Plantilla_Botón_1" at 1,715 size 130x53; TextOff 'PRINCIPAL'
      on Click: ActivateScreen("eProC - Principal", 0)
   Button "Template_Plantilla_Bouton_2" at 1085,715 size 193x53; TextOff 'ALARMAS / DEFAUT'
      on Press: ActivateScreen("eProC - Alarmas", 0)
      Visibility <- "DB_OP.P_DEFAUT"
   Button "Botón_6" at 374,621 size 88x33; TextOff 'Cerrar'
      on Press: SetTag("DB_OP.RC1", 52); SetBit("DB_OP.OP_SELMANU1")
      Visibility <- "MANU"
      Appearance <- "DB_OP.RC1"
   Button "Botón_7" at 374,578 size 88x33; TextOff 'Abrir'
      on Press: SetTag("DB_OP.RC1", 53); SetBit("DB_OP.OP_SELMANU1")
      Visibility <- "MANU"
      Appearance <- "DB_OP.RC1"
   Button "Botón_11" at 475,622 size 88x33; TextOff 'Freno'
      on Press: SetTag("DB_OP.RC1", 54); SetBit("DB_OP.OP_SELMANU1")
      Visibility <- "MANU"
      Appearance <- "DB_OP.RC1"
   Button "Botón_1" at 1002,622 size 88x33; TextOff 'Retroceso'
      on Press: SetTag("DB_OP.RC1", 55); SetBit("DB_OP.OP_SELMANU1")
      Visibility <- "MANU"
      Appearance <- "DB_OP.RC1"
   Button "Botón_2" at 1002,579 size 88x33; TextOff 'Avance'
      on Press: SetTag("DB_OP.RC1", 56); SetBit("DB_OP.OP_SELMANU1")
      Visibility <- "MANU"
      Appearance <- "DB_OP.RC1"
   TextField "Campo de texto_118" at 63,178 size 17x18; Text 'F1'
   IOField "Champ E/S_110" at 103,175 size 51x25; FormatPattern s999999
      Appearance <- "Perfiladores\Perfilador.PresenciaPieza"
      ProcessValue <- "Perfiladores\Perfilador.F1"
   IOField "Champ E/S_111" at 103,195 size 51x25; FormatPattern s999999
      Appearance <- "Perfiladores\Perfilador.PresenciaPieza"
      ProcessValue <- "Perfiladores\Perfilador.F2"
   IOField "Champ E/S_112" at 103,216 size 51x24; FormatPattern s999999
      Appearance <- "Perfiladores\Perfilador.PresenciaPieza"
      ProcessValue <- "Perfiladores\Perfilador.F3"
   IOField "Champ E/S_113" at 103,235 size 51x25; FormatPattern s999999
      Appearance <- "Perfiladores\Perfilador.PresenciaPieza"
      ProcessValue <- "Perfiladores\Perfilador.F4"
   TextField "Campo de texto_119" at 63,197 size 17x18; Text 'F2'
   TextField "Campo de texto_120" at 63,217 size 17x18; Text 'F3'
   TextField "Campo de texto_121" at 63,237 size 17x18; Text 'F4'
   TextField "Campo de texto_122" at 63,258 size 35x18; Text 'PL1-1'
   IOField "Champ E/S_114" at 103,255 size 51x25; FormatPattern s999999
      Appearance <- "Perfiladores\Perfilador.PresenciaPieza"
      ProcessValue <- "Perfiladores\Perfilador.PL1_1"
   IOField "Champ E/S_115" at 103,275 size 51x25; FormatPattern s999999
      Appearance <- "Perfiladores\Perfilador.PresenciaPieza"
      ProcessValue <- "Perfiladores\Perfilador.PL1_2"
   IOField "Champ E/S_116" at 103,296 size 51x24; FormatPattern s999999
      Appearance <- "Perfiladores\Perfilador.PresenciaPieza"
      ProcessValue <- "Perfiladores\Perfilador.PL2_1"
   IOField "Champ E/S_117" at 103,315 size 51x25; FormatPattern s999999
      Appearance <- "Perfiladores\Perfilador.PresenciaPieza"
      ProcessValue <- "Perfiladores\Perfilador.PL2_2"
   TextField "Campo de texto_123" at 63,278 size 35x18; Text 'PL1-2'
   TextField "Campo de texto_124" at 63,299 size 35x18; Text 'PL2-1'
   TextField "Campo de texto_125" at 63,318 size 35x18; Text 'PL2-2'

screen "eProC - 04 Cinta" 1280x768, template "Template"
   GraphicIOField "Campo ES gráfico_1" at 298,222 size 647x180; PictureList "Grupo 2 - Cinta"
      ProcessValue <- "Alarma_Cinta"
   Rectangle "Rectángulo_1" at 357,547 size 134x128
      Visibility <- "MANU"
   Rectangle "Rectángulo_2" at 986,116 size 118x128
      Visibility <- "MANU"
   Rectangle "Rectángulo_3" at 986,116 size 118x29
      Visibility <- "MANU"
   TextField "Campo de texto_1" at 1012,120 size 31x18; Text 'Cinta'
      Visibility <- "MANU"
   Rectangle "Rectángulo_7" at 357,531 size 134x29
      Visibility <- "MANU"
   TextField "Campo de texto_12" at 368,535 size 108x18; Text 'Ajuste Profundidad'
      Visibility <- "MANU"
   Circle "Cercle_1" at 333,248 size 12x12
      Appearance <- "27S4"
   Circle "Cercle_14" at 917,220 size 12x12
      Appearance <- "29S1"
   Circle "Cercle_15" at 917,234 size 12x12
      Appearance <- "29S2"
   Circle "Cercle_11" at 867,263 size 12x12
      Appearance <- "25S2"
   Circle "Cercle" at 927,268 size 12x12
      Appearance <- "29S3"
   TextField "Campo de texto_22" at 379,82 size 219x22; Text '27S4 - Chapa en Salida Perfilador'
   TextField "Campo de texto_23" at 632,433 size 213x22; Text 'M07 - Motor Ajuste Profundidad'
   TextField "Campo de texto_24" at 657,384 size 151x22; Text '25S2 - Bajar Velocidad'
   TextField "Campo de texto_25" at 992,311 size 269x22; Text '29S3 - Presencia de Chapa en Formador'
   TextField "Campo de texto_31" at 592,192 size 200x22; Text 'M08 - Motor Transporte Cinta'
   TextField "Campo de texto_32" at 643,128 size 172x22; Text '29S1 - Avance Bloqueado'
   TextField "Campo de texto_33" at 623,162 size 196x22; Text '29S2 - Avance Desbloqueado'
   Polygon "Polígono_4" at 356,247 size 472x69
      Visibility <- "Cinta\Cinta.PresenciaPieza"
   TextField "Campo de texto_113" at 59,77 size 31x18; Text 'Cinta'
   TextField "Campo de texto_114" at 59,99 size 12x18; Text 'A'
   IOField "Champ E/S_106" at 98,95 size 53x25; FormatPattern 9999999
      Appearance <- "Cinta\Cinta.PresenciaPieza"
      ProcessValue <- "Cinta\Cinta.A"
   IOField "Champ E/S_107" at 98,115 size 53x25; FormatPattern 9999999
      Appearance <- "Cinta\Cinta.PresenciaPieza"
      ProcessValue <- "Cinta\Cinta.B"
   IOField "Champ E/S_108" at 98,136 size 53x24; FormatPattern 9999999
      Appearance <- "Cinta\Cinta.PresenciaPieza"
      ProcessValue <- "Cinta\Cinta.C"
   IOField "Champ E/S_109" at 98,155 size 53x25; FormatPattern 9999999
      Appearance <- "Cinta\Cinta.PresenciaPieza"
      ProcessValue <- "Cinta\Cinta.D"
   TextField "Campo de texto_115" at 59,117 size 11x18; Text 'B'
   TextField "Campo de texto_116" at 59,137 size 11x18; Text 'C'
   TextField "Campo de texto_117" at 59,157 size 12x18; Text 'D'
   Button "Botón_14" at 43,40 size 126x33; TextOff 'Borrar Pieza'
      on Click: ResetBit("Cinta\Cinta.PresenciaPieza")
      Visibility <- "Cinta\Cinta.PresenciaPieza"
   Rectangle "Rectángulo_4" at 1114,116 size 118x128
      Visibility <- "MANU"
   Rectangle "Rectángulo_5" at 1114,116 size 118x29
      Visibility <- "MANU"
   TextField "Campo de texto_2" at 1140,120 size 33x18; Text 'Tope'
      Visibility <- "MANU"
   Button "Template_Plantilla_Botón_3" at 1,688 size 130x29; TextOff 'CINTA'
   Button "Plantilla_Botón_1" at 1,715 size 130x53; TextOff 'PRINCIPAL'
      on Click: ActivateScreen("eProC - Principal", 0)
   Button "Template_Plantilla_Bouton_2" at 1085,715 size 193x53; TextOff 'ALARMAS / DEFAUT'
      on Press: ActivateScreen("eProC - Alarmas", 0)
      Visibility <- "DB_OP.P_DEFAUT"
   Button "Botón_6" at 374,577 size 96x33; TextOff 'Avance'
      on Press: SetTag("DB_OP.RC1", 38); SetBit("DB_OP.OP_SELMANU1")
      Visibility <- "MANU"
      Appearance <- "DB_OP.RC1"
   Button "Botón_7" at 374,617 size 96x33; TextOff 'Retroceso'
      on Press: SetTag("DB_OP.RC1", 39); SetBit("DB_OP.OP_SELMANU1")
      Visibility <- "MANU"
      Appearance <- "DB_OP.RC1"
   Button "Botón_4" at 1000,159 size 88x33; TextOff 'Avance'
      on Press: SetTag("DB_OP.RC2", 91); SetBit("DB_OP.OP_SELMANU2")
      Visibility <- "MANU"
      Appearance <- "DB_OP.RC2"
   Button "Botón_5" at 1000,196 size 88x33; TextOff 'Retroceso'
      on Press: SetTag("DB_OP.RC2", 92); SetBit("DB_OP.OP_SELMANU2")
      Visibility <- "MANU"
      Appearance <- "DB_OP.RC2"
   Button "Botón_32" at 1127,196 size 94x33; TextOff 'Bajar Tope'
      on Press: SetTag("DB_OP.RC2", 36); SetBit("DB_OP.OP_SELMANU2")
      Visibility <- "MANU"
      Appearance <- "DB_OP.RC2"
   Button "Botón_33" at 1127,158 size 94x33; TextOff 'Subir Tope'
      on Press: SetTag("DB_OP.RC2", 35); SetBit("DB_OP.OP_SELMANU2")
      Visibility <- "MANU"
      Appearance <- "DB_OP.RC2"
   TextField "Campo de texto_150" at 61,178 size 17x18; Text 'F1'
   IOField "Champ E/S_142" at 101,175 size 51x25; FormatPattern s999999
      Appearance <- "Cinta\Cinta.PresenciaPieza"
      ProcessValue <- "Cinta\Cinta.F1"
   IOField "Champ E/S_143" at 101,195 size 51x25; FormatPattern s999999
      Appearance <- "Cinta\Cinta.PresenciaPieza"
      ProcessValue <- "Cinta\Cinta.F2"
   IOField "Champ E/S_144" at 101,216 size 51x24; FormatPattern s999999
      Appearance <- "Cinta\Cinta.PresenciaPieza"
      ProcessValue <- "Cinta\Cinta.F3"
   IOField "Champ E/S_145" at 101,235 size 51x25; FormatPattern s999999
      Appearance <- "Cinta\Cinta.PresenciaPieza"
      ProcessValue <- "Cinta\Cinta.F4"
   TextField "Campo de texto_151" at 61,197 size 17x18; Text 'F2'
   TextField "Campo de texto_152" at 61,217 size 17x18; Text 'F3'
   TextField "Campo de texto_153" at 61,237 size 17x18; Text 'F4'
   TextField "Campo de texto_154" at 61,258 size 35x18; Text 'PL1-1'
   IOField "Champ E/S_146" at 101,255 size 51x25; FormatPattern s999999
      Appearance <- "Cinta\Cinta.PresenciaPieza"
      ProcessValue <- "Cinta\Cinta.PL1_1"
   IOField "Champ E/S_147" at 101,275 size 51x25; FormatPattern s999999
      Appearance <- "Cinta\Cinta.PresenciaPieza"
      ProcessValue <- "Cinta\Cinta.PL1_2"
   IOField "Champ E/S_148" at 101,296 size 51x24; FormatPattern s999999
      Appearance <- "Cinta\Cinta.PresenciaPieza"
      ProcessValue <- "Cinta\Cinta.PL2_1"
   IOField "Champ E/S_149" at 101,315 size 51x25; FormatPattern s999999
      Appearance <- "Cinta\Cinta.PresenciaPieza"
      ProcessValue <- "Cinta\Cinta.PL2_2"
   TextField "Campo de texto_155" at 61,278 size 35x18; Text 'PL1-2'
   TextField "Campo de texto_156" at 61,299 size 35x18; Text 'PL2-1'
   TextField "Campo de texto_157" at 61,318 size 35x18; Text 'PL2-2'